   "Carrier_22_First_Duplicate_Carrier_Position" AT %QD1468 : DWord;
   "Carrier_22_Second_Duplicate_Carrier_Position" AT %QD1472 : DWord;
   "Carrier_22_CommandWord" AT %QW1476 : Word;
   "Carrier_22_Heartbeat" AT %Q1476.0 : Bool;
   "Carrier_22_Drive_Forward_Command" AT %Q1476.1 : Bool;
   "Carrier_22_Fault_Reset" AT %Q1476.2 : Bool;
   "Carrier_22_At_Command_Position" AT %Q1476.3 : Bool;
   "Carrier_22_Duplicate_Carrier_Fault" AT %Q1476.4 : Bool;
   "Carrier_22_Motion_On_Fault" AT %Q1476.5 : Bool;
   "Carrier_22_Motion_Off_Fault" AT %Q1476.6 : Bool;
   "Carrier_22_Carrier_Spacing_Fault" AT %Q1476.7 : Bool;
   "Carrier_23_Carrier_In_Zone" AT %QW1500 : Word;
   "Carrier_23_Carrier_Number_Echo" AT %QW1502 : Word;
   "Carrier_23_Carrier_Position_Echo" AT %QD1504 : DWord;
   "Carrier_23_Next_Carrier_Number" AT %QW1508 : Word;
   "Carrier_23_Next_Stop_Position" AT %QD1510 : DWord;
   "Carrier_23_Drive_Command_Speed" AT %QW1514 : Word;
   "Carrier_23_Duplicate_Carrier_Number" AT %QW1516 : Word;
   "Carrier_23_First_Duplicate_Carrier_Position" AT %QD1518 : DWord;
   "Carrier_23_Second_Duplicate_Carrier_Position" AT %QD1522 : DWord;
   "Carrier_23_CommandWord" AT %QW1526 : Word;
   "Carrier_23_Heartbeat" AT %Q1526.0 : Bool;
   "Carrier_23_Drive_Forward_Command" AT %Q1526.1 : Bool;
   "Carrier_23_Fault_Reset" AT %Q1526.2 : Bool;
   "Carrier_23_At_Command_Position" AT %Q1526.3 : Bool;
   "Carrier_23_Duplicate_Carrier_Fault" AT %Q1526.4 : Bool;
   "Carrier_23_Motion_On_Fault" AT %Q1526.5 : Bool;
   "Carrier_23_Motion_Off_Fault" AT %Q1526.6 : Bool;
   "Carrier_23_Carrier_Spacing_Fault" AT %Q1526.7 : Bool;
   "Carrier_24_Carrier_In_Zone" AT %QW1550 : Word;
   "Carrier_24_Carrier_Number_Echo" AT %QW1552 : Word;
   "Carrier_24_Carrier_Position_Echo" AT %QD1554 : DWord;
   "Carrier_24_Next_Carrier_Number" AT %QW1558 : Word;
   "Carrier_24_Next_Stop_Position" AT %QD1560 : DWord;
   "Carrier_24_Drive_Command_Speed" AT %QW1564 : Word;
   "Carrier_24_Duplicate_Carrier_Number" AT %QW1566 : Word;
   "Carrier_24_First_Duplicate_Carrier_Position" AT %QD1568 : DWord;
   "Carrier_24_Second_Duplicate_Carrier_Position" AT %QD1572 : DWord;
   "Carrier_24_CommandWord" AT %QW1576 : Word;
   "Carrier_24_Heartbeat" AT %Q1576.0 : Bool;
   "Carrier_24_Drive_Forward_Command" AT %Q1576.1 : Bool;
   "Carrier_24_Fault_Reset" AT %Q1576.2 : Bool;
   "Carrier_24_At_Command_Position" AT %Q1576.3 : Bool;
   "Carrier_24_Duplicate_Carrier_Fault" AT %Q1576.4 : Bool;
   "Carrier_24_Motion_On_Fault" AT %Q1576.5 : Bool;
   "Carrier_24_Motion_Off_Fault" AT %Q1576.6 : Bool;
   "Carrier_24_Carrier_Spacing_Fault" AT %Q1576.7 : Bool;
   "Carrier_25_Carrier_In_Zone" AT %QW1600 : Word;
   "Carrier_25_Carrier_Number_Echo" AT %QW1602 : Word;
   "Carrier_25_Carrier_Position_Echo" AT %QD1604 : DWord;
   "Carrier_25_Next_Carrier_Number" AT %QW1608 : Word;
   "Carrier_25_Next_Stop_Position" AT %QD1610 : DWord;
   "Carrier_25_Drive_Command_Speed" AT %QW1614 : Word;
   "Carrier_25_Duplicate_Carrier_Number" AT %QW1616 : Word;
   "Carrier_25_First_Duplicate_Carrier_Position" AT %QD1618 : DWord;
   "Carrier_25_Second_Duplicate_Carrier_Position" AT %QD1622 : DWord;
   "Carrier_25_CommandWord" AT %QW1626 : Word;
   "Carrier_25_Heartbeat" AT %Q1626.0 : Bool;
   "Carrier_25_Drive_Forward_Command" AT %Q1626.1 : Bool;
   "Carrier_25_Fault_Reset" AT %Q1626.2 : Bool;
   "Carrier_25_At_Command_Position" AT %Q1626.3 : Bool;
   "Carrier_25_Duplicate_Carrier_Fault" AT %Q1626.4 : Bool;
   "Carrier_25_Motion_On_Fault" AT %Q1626.5 : Bool;
   "Carrier_25_Motion_Off_Fault" AT %Q1626.6 : Bool;
   "Carrier_25_Carrier_Spacing_Fault" AT %Q1626.7 : Bool;
   "Carrier_26_Carrier_In_Zone" AT %QW1650 : Word;
   "Carrier_26_Carrier_Number_Echo" AT %QW1652 : Word;
   "Carrier_26_Carrier_Position_Echo" AT %QD1654 : DWord;
   "Carrier_26_Next_Carrier_Number" AT %QW1658 : Word;
   "Carrier_26_Next_Stop_Position" AT %QD1660 : DWord;
   "Carrier_26_Drive_Command_Speed" AT %QW1664 : Word;
   "Carrier_26_Duplicate_Carrier_Number" AT %QW1666 : Word;
   "Carrier_26_First_Duplicate_Carrier_Position" AT %QD1668 : DWord;
   "Carrier_26_Second_Duplicate_Carrier_Position" AT %QD1672 : DWord;
   "Carrier_26_CommandWord" AT %QW1676 : Word;
   "Carrier_26_Heartbeat" AT %Q1676.0 : Bool;
   "Carrier_26_Drive_Forward_Command" AT %Q1676.1 : Bool;
   "Carrier_26_Fault_Reset" AT %Q1676.2 : Bool;
   "Carrier_26_At_Command_Position" AT %Q1676.3 : Bool;
   "Carrier_26_Duplicate_Carrier_Fault" AT %Q1676.4 : Bool;
   "Carrier_26_Motion_On_Fault" AT %Q1676.5 : Bool;
   "Carrier_26_Motion_Off_Fault" AT %Q1676.6 : Bool;
   "Carrier_26_Carrier_Spacing_Fault" AT %Q1676.7 : Bool;
   "Carrier_27_Carrier_In_Zone" AT %QW1700 : Word;
   "Carrier_27_Carrier_Number_Echo" AT %QW1702 : Word;
   "Carrier_27_Carrier_Position_Echo" AT %QD1704 : DWord;
   "Carrier_27_Next_Carrier_Number" AT %QW1708 : Word;
   "Carrier_27_Next_Stop_Position" AT %QD1710 : DWord;
   "Carrier_27_Drive_Command_Speed" AT %QW1714 : Word;
   "Carrier_27_Duplicate_Carrier_Number" AT %QW1716 : Word;
   "Carrier_27_First_Duplicate_Carrier_Position" AT %QD1718 : DWord;
   "Carrier_27_Second_Duplicate_Carrier_Position" AT %QD1722 : DWord;
   "Carrier_27_CommandWord" AT %QW1726 : Word;
   "Carrier_27_Heartbeat" AT %Q1726.0 : Bool;
   "Carrier_27_Drive_Forward_Command" AT %Q1726.1 : Bool;
   "Carrier_27_Fault_Reset" AT %Q1726.2 : Bool;
   "Carrier_27_At_Command_Position" AT %Q1726.3 : Bool;
   "Carrier_27_Duplicate_Carrier_Fault" AT %Q1726.4 : Bool;
   "Carrier_27_Motion_On_Fault" AT %Q1726.5 : Bool;
   "Carrier_27_Motion_Off_Fault" AT %Q1726.6 : Bool;
   "Carrier_27_Carrier_Spacing_Fault" AT %Q1726.7 : Bool;
   "Carrier_28_Carrier_In_Zone" AT %QW1750 : Word;
   "Carrier_28_Carrier_Number_Echo" AT %QW1752 : Word;
   "Carrier_28_Carrier_Position_Echo" AT %QD1754 : DWord;
   "Carrier_28_Next_Carrier_Number" AT %QW1758 : Word;
   "Carrier_28_Next_Stop_Position" AT %QD1760 : DWord;
   "Carrier_28_Drive_Command_Speed" AT %QW1764 : Word;
   "Carrier_28_Duplicate_Carrier_Number" AT %QW1766 : Word;
   "Carrier_28_First_Duplicate_Carrier_Position" AT %QD1768 : DWord;
   "Carrier_28_Second_Duplicate_Carrier_Position" AT %QD1772 : DWord;
   "Carrier_28_CommandWord" AT %QW1776 : Word;
   "Carrier_28_Heartbeat" AT %Q1776.0 : Bool;
   "Carrier_28_Drive_Forward_Command" AT %Q1776.1 : Bool;
   "Carrier_28_Fault_Reset" AT %Q1776.2 : Bool;
   "Carrier_28_At_Command_Position" AT %Q1776.3 : Bool;
   "Carrier_28_Duplicate_Carrier_Fault" AT %Q1776.4 : Bool;
   "Carrier_28_Motion_On_Fault" AT %Q1776.5 : Bool;
   "Carrier_28_Motion_Off_Fault" AT %Q1776.6 : Bool;
   "Carrier_28_Carrier_Spacing_Fault" AT %Q1776.7 : Bool;
   "Carrier_29_Carrier_In_Zone" AT %QW1800 : Word;
   "Carrier_29_Carrier_Number_Echo" AT %QW1802 : Word;
   "Carrier_29_Carrier_Position_Echo" AT %QD1804 : DWord;
   "Carrier_29_Next_Carrier_Number" AT %QW1808 : Word;
   "Carrier_29_Next_Stop_Position" AT %QD1810 : DWord;
   "Carrier_29_Drive_Command_Speed" AT %QW1814 : Word;
   "Carrier_29_Duplicate_Carrier_Number" AT %QW1816 : Word;
   "Carrier_29_First_Duplicate_Carrier_Position" AT %QD1818 : DWord;
   "Carrier_29_Second_Duplicate_Carrier_Position" AT %QD1822 : DWord;
   "Carrier_29_CommandWord" AT %QW1826 : Word;
   "Carrier_29_Heartbeat" AT %Q1826.0 : Bool;
   "Carrier_29_Drive_Forward_Command" AT %Q1826.1 : Bool;
   "Carrier_29_Fault_Reset" AT %Q1826.2 : Bool;
   "Carrier_29_At_Command_Position" AT %Q1826.3 : Bool;
   "Carrier_29_Duplicate_Carrier_Fault" AT %Q1826.4 : Bool;
   "Carrier_29_Motion_On_Fault" AT %Q1826.5 : Bool;
   "Carrier_29_Motion_Off_Fault" AT %Q1826.6 : Bool;
   "Carrier_29_Carrier_Spacing_Fault" AT %Q1826.7 : Bool;
   "Carrier_30_Carrier_In_Zone" AT %QW1850 : Word;
   "Carrier_30_Carrier_Number_Echo" AT %QW1852 : Word;
   "Carrier_30_Carrier_Position_Echo" AT %QD1854 : DWord;
   "Carrier_30_Next_Carrier_Number" AT %QW1858 : Word;
   "Carrier_30_Next_Stop_Position" AT %QD1860 : DWord;
   "Carrier_30_Drive_Command_Speed" AT %QW1864 : Word;
   "Carrier_30_Duplicate_Carrier_Number" AT %QW1866 : Word;
   "Carrier_30_First_Duplicate_Carrier_Position" AT %QD1868 : DWord;
   "Carrier_30_Second_Duplicate_Carrier_Position" AT %QD1872 : DWord;
   "Carrier_30_CommandWord" AT %QW1876 : Word;
   "Carrier_30_Heartbeat" AT %Q1876.0 : Bool;
   "Carrier_30_Drive_Forward_Command" AT %Q1876.1 : Bool;
   "Carrier_30_Fault_Reset" AT %Q1876.2 : Bool;
   "Carrier_30_At_Command_Position" AT %Q1876.3 : Bool;
   "Carrier_30_Duplicate_Carrier_Fault" AT %Q1876.4 : Bool;
   "Carrier_30_Motion_On_Fault" AT %Q1876.5 : Bool;
   "Carrier_30_Motion_Off_Fault" AT %Q1876.6 : Bool;
   "Carrier_30_Carrier_Spacing_Fault" AT %Q1876.7 : Bool;
   "Carrier_31_Carrier_In_Zone" AT %QW1900 : Word;
   "Carrier_31_Carrier_Number_Echo" AT %QW1902 : Word;
   "Carrier_31_Carrier_Position_Echo" AT %QD1904 : DWord;
   "Carrier_31_Next_Carrier_Number" AT %QW1908 : Word;
   "Carrier_31_Next_Stop_Position" AT %QD1910 : DWord;
   "Carrier_31_Drive_Command_Speed" AT %QW1914 : Word;
   "Carrier_31_Duplicate_Carrier_Number" AT %QW1916 : Word;
   "Carrier_31_First_Duplicate_Carrier_Position" AT %QD1918 : DWord;
   "Carrier_31_Second_Duplicate_Carrier_Position" AT %QD1922 : DWord;
   "Carrier_31_CommandWord" AT %QW1926 : Word;
   "Carrier_31_Heartbeat" AT %Q1926.0 : Bool;
   "Carrier_31_Drive_Forward_Command" AT %Q1926.1 : Bool;
   "Carrier_31_Fault_Reset" AT %Q1926.2 : Bool;
   "Carrier_31_At_Command_Position" AT %Q1926.3 : Bool;
   "Carrier_31_Duplicate_Carrier_Fault" AT %Q1926.4 : Bool;
   "Carrier_31_Motion_On_Fault" AT %Q1926.5 : Bool;
   "Carrier_31_Motion_Off_Fault" AT %Q1926.6 : Bool;
   "Carrier_31_Carrier_Spacing_Fault" AT %Q1926.7 : Bool;
   "Carrier_32_Carrier_In_Zone" AT %QW1950 : Word;
   "Carrier_32_Carrier_Number_Echo" AT %QW1952 : Word;
   "Carrier_32_Carrier_Position_Echo" AT %QD1954 : DWord;
   "Carrier_32_Next_Carrier_Number" AT %QW1958 : Word;
   "Carrier_32_Next_Stop_Position" AT %QD1960 : DWord;
   "Carrier_32_Drive_Command_Speed" AT %QW1964 : Word;
   "Carrier_32_Duplicate_Carrier_Number" AT %QW1966 : Word;
   "Carrier_32_First_Duplicate_Carrier_Position" AT %QD1968 : DWord;
   "Carrier_32_Second_Duplicate_Carrier_Position" AT %QD1972 : DWord;
   "Carrier_32_CommandWord" AT %QW1976 : Word;
   "Carrier_32_Heartbeat" AT %Q1976.0 : Bool;
   "Carrier_32_Drive_Forward_Command" AT %Q1976.1 : Bool;
   "Carrier_32_Fault_Reset" AT %Q1976.2 : Bool;
   "Carrier_32_At_Command_Position" AT %Q1976.3 : Bool;
   "Carrier_32_Duplicate_Carrier_Fault" AT %Q1976.4 : Bool;
   "Carrier_32_Motion_On_Fault" AT %Q1976.5 : Bool;
   "Carrier_32_Motion_Off_Fault" AT %Q1976.6 : Bool;
   "Carrier_32_Carrier_Spacing_Fault" AT %Q1976.7 : Bool;
   "Carrier_33_Carrier_In_Zone" AT %QW2000 : Word;
   "Carrier_33_Carrier_Number_Echo" AT %QW2002 : Word;
   "Carrier_33_Carrier_Position_Echo" AT %QD2004 : DWord;
   "Carrier_33_Next_Carrier_Number" AT %QW2008 : Word;
   "Carrier_33_Next_Stop_Position" AT %QD2010 : DWord;
   "Carrier_33_Drive_Command_Speed" AT %QW2014 : Word;
   "Carrier_33_Duplicate_Carrier_Number" AT %QW2016 : Word;
   "Carrier_33_First_Duplicate_Carrier_Position" AT %QD2018 : DWord;
   "Carrier_33_Second_Duplicate_Carrier_Position" AT %QD2022 : DWord;
   "Carrier_33_CommandWord" AT %QW2026 : Word;
   "Carrier_33_Heartbeat" AT %Q2026.0 : Bool;
   "Carrier_33_Drive_Forward_Command" AT %Q2026.1 : Bool;
   "Carrier_33_Fault_Reset" AT %Q2026.2 : Bool;
   "Carrier_33_At_Command_Position" AT %Q2026.3 : Bool;
   "Carrier_33_Duplicate_Carrier_Fault" AT %Q2026.4 : Bool;
   "Carrier_33_Motion_On_Fault" AT %Q2026.5 : Bool;
   "Carrier_33_Motion_Off_Fault" AT %Q2026.6 : Bool;
   "Carrier_33_Carrier_Spacing_Fault" AT %Q2026.7 : Bool;
   "Carrier_34_Carrier_In_Zone" AT %QW2050 : Word;
   "Carrier_34_Carrier_Number_Echo" AT %QW2052 : Word;
   "Carrier_34_Carrier_Position_Echo" AT %QD2054 : DWord;
   "Carrier_34_Next_Carrier_Number" AT %QW2058 : Word;
   "Carrier_34_Next_Stop_Position" AT %QD2060 : DWord;
   "Carrier_34_Drive_Command_Speed" AT %QW2064 : Word;
   "Carrier_34_Duplicate_Carrier_Number" AT %QW2066 : Word;
   "Carrier_34_First_Duplicate_Carrier_Position" AT %QD2068 : DWord;
   "Carrier_34_Second_Duplicate_Carrier_Position" AT %QD2072 : DWord;
   "Carrier_34_CommandWord" AT %QW2076 : Word;
   "Carrier_34_Heartbeat" AT %Q2076.0 : Bool;
   "Carrier_34_Drive_Forward_Command" AT %Q2076.1 : Bool;
   "Carrier_34_Fault_Reset" AT %Q2076.2 : Bool;
   "Carrier_34_At_Command_Position" AT %Q2076.3 : Bool;
   "Carrier_34_Duplicate_Carrier_Fault" AT %Q2076.4 : Bool;
   "Carrier_34_Motion_On_Fault" AT %Q2076.5 : Bool;
   "Carrier_34_Motion_Off_Fault" AT %Q2076.6 : Bool;
   "Carrier_34_Carrier_Spacing_Fault" AT %Q2076.7 : Bool;
   "Carrier_35_Carrier_In_Zone" AT %QW2100 : Word;
   "Carrier_35_Carrier_Number_Echo" AT %QW2102 : Word;
   "Carrier_35_Carrier_Position_Echo" AT %QD2104 : DWord;
   "Carrier_35_Next_Carrier_Number" AT %QW2108 : Word;
   "Carrier_35_Next_Stop_Position" AT %QD2110 : DWord;
   "Carrier_35_Drive_Command_Speed" AT %QW2114 : Word;
   "Carrier_35_Duplicate_Carrier_Number" AT %QW2116 : Word;
   "Carrier_35_First_Duplicate_Carrier_Position" AT %QD2118 : DWord;
   "Carrier_35_Second_Duplicate_Carrier_Position" AT %QD2122 : DWord;
   "Carrier_35_CommandWord" AT %QW2126 : Word;
   "Carrier_35_Heartbeat" AT %Q2126.0 : Bool;
   "Carrier_35_Drive_Forward_Command" AT %Q2126.1 : Bool;
   "Carrier_35_Fault_Reset" AT %Q2126.2 : Bool;
   "Carrier_35_At_Command_Position" AT %Q2126.3 : Bool;
   "Carrier_35_Duplicate_Carrier_Fault" AT %Q2126.4 : Bool;
   "Carrier_35_Motion_On_Fault" AT %Q2126.5 : Bool;
   "Carrier_35_Motion_Off_Fault" AT %Q2126.6 : Bool;
   "Carrier_35_Carrier_Spacing_Fault" AT %Q2126.7 : Bool;
   "Carrier_36_Carrier_In_Zone" AT %QW2150 : Word;
   "Carrier_36_Carrier_Number_Echo" AT %QW2152 : Word;
   "Carrier_36_Carrier_Position_Echo" AT %QD2154 : DWord;
   "Carrier_36_Next_Carrier_Number" AT %QW2158 : Word;
   "Carrier_36_Next_Stop_Position" AT %QD2160 : DWord;
   "Carrier_36_Drive_Command_Speed" AT %QW2164 : Word;
   "Carrier_36_Duplicate_Carrier_Number" AT %QW2166 : Word;
   "Carrier_36_First_Duplicate_Carrier_Position" AT %QD2168 : DWord;
   "Carrier_36_Second_Duplicate_Carrier_Position" AT %QD2172 : DWord;
   "Carrier_36_CommandWord" AT %QW2176 : Word;
   "Carrier_36_Heartbeat" AT %Q2176.0 : Bool;
   "Carrier_36_Drive_Forward_Command" AT %Q2176.1 : Bool;
   "Carrier_36_Fault_Reset" AT %Q2176.2 : Bool;
   "Carrier_36_At_Command_Position" AT %Q2176.3 : Bool;
   "Carrier_36_Duplicate_Carrier_Fault" AT %Q2176.4 : Bool;
   "Carrier_36_Motion_On_Fault" AT %Q2176.5 : Bool;
   "Carrier_36_Motion_Off_Fault" AT %Q2176.6 : Bool;
   "Carrier_36_Carrier_Spacing_Fault" AT %Q2176.7 : Bool;
   "Carrier_37_Carrier_In_Zone" AT %QW2200 : Word;
   "Carrier_37_Carrier_Number_Echo" AT %QW2202 : Word;
   "Carrier_37_Carrier_Position_Echo" AT %QD2204 : DWord;
   "Carrier_37_Next_Carrier_Number" AT %QW2208 : Word;
   "Carrier_37_Next_Stop_Position" AT %QD2210 : DWord;
   "Carrier_37_Drive_Command_Speed" AT %QW2214 : Word;
   "Carrier_37_Duplicate_Carrier_Number" AT %QW2216 : Word;
   "Carrier_37_First_Duplicate_Carrier_Position" AT %QD2218 : DWord;
   "Carrier_37_Second_Duplicate_Carrier_Position" AT %QD2222 : DWord;
   "Carrier_37_CommandWord" AT %QW2226 : Word;
   "Carrier_37_Heartbeat" AT %Q2226.0 : Bool;
   "Carrier_37_Drive_Forward_Command" AT %Q2226.1 : Bool;
   "Carrier_37_Fault_Reset" AT %Q2226.2 : Bool;
   "Carrier_37_At_Command_Position" AT %Q2226.3 : Bool;
   "Carrier_37_Duplicate_Carrier_Fault" AT %Q2226.4 : Bool;
   "Carrier_37_Motion_On_Fault" AT %Q2226.5 : Bool;
   "Carrier_37_Motion_Off_Fault" AT %Q2226.6 : Bool;
   "Carrier_37_Carrier_Spacing_Fault" AT %Q2226.7 : Bool;
   "Carrier_38_Carrier_In_Zone" AT %QW2250 : Word;
   "Carrier_38_Carrier_Number_Echo" AT %QW2252 : Word;
   "Carrier_38_Carrier_Position_Echo" AT %QD2254 : DWord;
   "Carrier_38_Next_Carrier_Number" AT %QW2258 : Word;
   "Carrier_38_Next_Stop_Position" AT %QD2260 : DWord;
   "Carrier_38_Drive_Command_Speed" AT %QW2264 : Word;
   "Carrier_38_Duplicate_Carrier_Number" AT %QW2266 : Word;
   "Carrier_38_First_Duplicate_Carrier_Position" AT %QD2268 : DWord;
   "Carrier_38_Second_Duplicate_Carrier_Position" AT %QD2272 : DWord;
   "Carrier_38_CommandWord" AT %QW2276 : Word;
   "Carrier_38_Heartbeat" AT %Q2276.0 : Bool;
   "Carrier_38_Drive_Forward_Command" AT %Q2276.1 : Bool;
   "Carrier_38_Fault_Reset" AT %Q2276.2 : Bool;
   "Carrier_38_At_Command_Position" AT %Q2276.3 : Bool;
   "Carrier_38_Duplicate_Carrier_Fault" AT %Q2276.4 : Bool;
   "Carrier_38_Motion_On_Fault" AT %Q2276.5 : Bool;
   "Carrier_38_Motion_Off_Fault" AT %Q2276.6 : Bool;
   "Carrier_38_Carrier_Spacing_Fault" AT %Q2276.7 : Bool;
   "Carrier_39_Carrier_In_Zone" AT %QW2300 : Word;
   "Carrier_39_Carrier_Number_Echo" AT %QW2302 : Word;
   "Carrier_39_Carrier_Position_Echo" AT %QD2304 : DWord;
   "Carrier_39_Next_Carrier_Number" AT %QW2308 : Word;
   "Carrier_39_Next_Stop_Position" AT %QD2310 : DWord;
   "Carrier_39_Drive_Command_Speed" AT %QW2314 : Word;
   "Carrier_39_Duplicate_Carrier_Number" AT %QW2316 : Word;
   "Carrier_39_First_Duplicate_Carrier_Position" AT %QD2318 : DWord;
   "Carrier_39_Second_Duplicate_Carrier_Position" AT %QD2322 : DWord;
   "Carrier_39_CommandWord" AT %QW2326 : Word;
   "Carrier_39_Heartbeat" AT %Q2326.0 : Bool;
   "Carrier_39_Drive_Forward_Command" AT %Q2326.1 : Bool;
   "Carrier_39_Fault_Reset" AT %Q2326.2 : Bool;
   "Carrier_39_At_Command_Position" AT %Q2326.3 : Bool;
   "Carrier_39_Duplicate_Carrier_Fault" AT %Q2326.4 : Bool;
   "Carrier_39_Motion_On_Fault" AT %Q2326.5 : Bool;
   "Carrier_39_Motion_Off_Fault" AT %Q2326.6 : Bool;
   "Carrier_39_Carrier_Spacing_Fault" AT %Q2326.7 : Bool;
   "Carrier_40_Carrier_In_Zone" AT %QW2350 : Word;
   "Carrier_40_Carrier_Number_Echo" AT %QW2352 : Word;
   "Carrier_40_Carrier_Position_Echo" AT %QD2354 : DWord;
   "Carrier_40_Next_Carrier_Number" AT %QW2358 : Word;
   "Carrier_40_Next_Stop_Position" AT %QD2360 : DWord;
   "Carrier_40_Drive_Command_Speed" AT %QW2364 : Word;
   "Carrier_40_Duplicate_Carrier_Number" AT %QW2366 : Word;
   "Carrier_40_First_Duplicate_Carrier_Position" AT %QD2368 : DWord;
   "Carrier_40_Second_Duplicate_Carrier_Position" AT %QD2372 : DWord;
   "Carrier_40_CommandWord" AT %QW2376 : Word;
   "Carrier_40_Heartbeat" AT %Q2376.0 : Bool;
   "Carrier_40_Drive_Forward_Command" AT %Q2376.1 : Bool;
   "Carrier_40_Fault_Reset" AT %Q2376.2 : Bool;
   "Carrier_40_At_Command_Position" AT %Q2376.3 : Bool;
   "Carrier_40_Duplicate_Carrier_Fault" AT %Q2376.4 : Bool;
   "Carrier_40_Motion_On_Fault" AT %Q2376.5 : Bool;
   "Carrier_40_Motion_Off_Fault" AT %Q2376.6 : Bool;
   "Carrier_40_Carrier_Spacing_Fault" AT %Q2376.7 : Bool;
   "Carrier_41_Carrier_In_Zone" AT %QW2400 : Word;
   "Carrier_41_Carrier_Number_Echo" AT %QW2402 : Word;
   "Carrier_41_Carrier_Position_Echo" AT %QD2404 : DWord;
   "Carrier_41_Next_Carrier_Number" AT %QW2408 : Word;
   "Carrier_41_Next_Stop_Position" AT %QD2410 : DWord;
   "Carrier_41_Drive_Command_Speed" AT %QW2414 : Word;
   "Carrier_41_Duplicate_Carrier_Number" AT %QW2416 : Word;
   "Carrier_41_First_Duplicate_Carrier_Position" AT %QD2418 : DWord;
   "Carrier_41_Second_Duplicate_Carrier_Position" AT %QD2422 : DWord;
   "Carrier_41_CommandWord" AT %QW2426 : Word;
   "Carrier_41_Heartbeat" AT %Q2426.0 : Bool;
   "Carrier_41_Drive_Forward_Command" AT %Q2426.1 : Bool;
   "Carrier_41_Fault_Reset" AT %Q2426.2 : Bool;
   "Carrier_41_At_Command_Position" AT %Q2426.3 : Bool;
   "Carrier_41_Duplicate_Carrier_Fault" AT %Q2426.4 : Bool;
   "Carrier_41_Motion_On_Fault" AT %Q2426.5 : Bool;
   "Carrier_41_Motion_Off_Fault" AT %Q2426.6 : Bool;
   "Carrier_41_Carrier_Spacing_Fault" AT %Q2426.7 : Bool;
   "Carrier_42_Carrier_In_Zone" AT %QW2450 : Word;
   "Carrier_42_Carrier_Number_Echo" AT %QW2452 : Word;
   "Carrier_42_Carrier_Position_Echo" AT %QD2454 : DWord;
   "Carrier_42_Next_Carrier_Number" AT %QW2458 : Word;
   "Carrier_42_Next_Stop_Position" AT %QD2460 : DWord;
   "Carrier_42_Drive_Command_Speed" AT %QW2464 : Word;
   "Carrier_42_Duplicate_Carrier_Number" AT %QW2466 : Word;
   "Carrier_42_First_Duplicate_Carrier_Position" AT %QD2468 : DWord;
   "Carrier_42_Second_Duplicate_Carrier_Position" AT %QD2472 : DWord;
   "Carrier_42_CommandWord" AT %QW2476 : Word;
   "Carrier_42_Heartbeat" AT %Q2476.0 : Bool;
   "Carrier_42_Drive_Forward_Command" AT %Q2476.1 : Bool;
   "Carrier_42_Fault_Reset" AT %Q2476.2 : Bool;
   "Carrier_42_At_Command_Position" AT %Q2476.3 : Bool;
   "Carrier_42_Duplicate_Carrier_Fault" AT %Q2476.4 : Bool;
   "Carrier_42_Motion_On_Fault" AT %Q2476.5 : Bool;
   "Carrier_42_Motion_Off_Fault" AT %Q2476.6 : Bool;
   "Carrier_42_Carrier_Spacing_Fault" AT %Q2476.7 : Bool;
   "Carrier_43_Carrier_In_Zone" AT %QW2500 : Word;
   "Carrier_43_Carrier_Number_Echo" AT %QW2502 : Word;
   "Carrier_43_Carrier_Position_Echo" AT %QD2504 : DWord;
   "Carrier_43_Next_Carrier_Number" AT %QW2508 : Word;
   "Carrier_43_Next_Stop_Position" AT %QD2510 : DWord;
   "Carrier_43_Drive_Command_Speed" AT %QW2514 : Word;
   "Carrier_43_Duplicate_Carrier_Number" AT %QW2516 : Word;
   "Carrier_43_First_Duplicate_Carrier_Position" AT %QD2518 : DWord;
   "Carrier_43_Second_Duplicate_Carrier_Position" AT %QD2522 : DWord;
   "Carrier_43_CommandWord" AT %QW2526 : Word;
   "Carrier_43_Heartbeat" AT %Q2526.0 : Bool;
   "Carrier_43_Drive_Forward_Command" AT %Q2526.1 : Bool;
   "Carrier_43_Fault_Reset" AT %Q2526.2 : Bool;
   "Carrier_43_At_Command_Position" AT %Q2526.3 : Bool;
   "Carrier_43_Duplicate_Carrier_Fault" AT %Q2526.4 : Bool;
   "Carrier_43_Motion_On_Fault" AT %Q2526.5 : Bool;
   "Carrier_43_Motion_Off_Fault" AT %Q2526.6 : Bool;
   "Carrier_43_Carrier_Spacing_Fault" AT %Q2526.7 : Bool;
   "Carrier_44_Carrier_In_Zone" AT %QW2550 : Word;
   "Carrier_44_Carrier_Number_Echo" AT %QW2552 : Word;
   "Carrier_44_Carrier_Position_Echo" AT %QD2554 : DWord;
   "Carrier_44_Next_Carrier_Number" AT %QW2558 : Word;
   "Carrier_44_Next_Stop_Position" AT %QD2560 : DWord;
   "Carrier_44_Drive_Command_Speed" AT %QW2564 : Word;
   "Carrier_44_Duplicate_Carrier_Number" AT %QW2566 : Word;
   "Carrier_44_First_Duplicate_Carrier_Position" AT %QD2568 : DWord;
   "Carrier_44_Second_Duplicate_Carrier_Position" AT %QD2572 : DWord;
   "Carrier_44_CommandWord" AT %QW2576 : Word;
   "Carrier_44_Heartbeat" AT %Q2576.0 : Bool;
   "Carrier_44_Drive_Forward_Command" AT %Q2576.1 : Bool;
   "Carrier_44_Fault_Reset" AT %Q2576.2 : Bool;
   "Carrier_44_At_Command_Position" AT %Q2576.3 : Bool;
   "Carrier_44_Duplicate_Carrier_Fault" AT %Q2576.4 : Bool;
   "Carrier_44_Motion_On_Fault" AT %Q2576.5 : Bool;
   "Carrier_44_Motion_Off_Fault" AT %Q2576.6 : Bool;
   "Carrier_44_Carrier_Spacing_Fault" AT %Q2576.7 : Bool;
   "Carrier_45_Carrier_In_Zone" AT %QW2600 : Word;
   "Carrier_45_Carrier_Number_Echo" AT %QW2602 : Word;
   "Carrier_45_Carrier_Position_Echo" AT %QD2604 : DWord;
   "Carrier_45_Next_Carrier_Number" AT %QW2608 : Word;
   "Carrier_45_Next_Stop_Position" AT %QD2610 : DWord;
   "Carrier_45_Drive_Command_Speed" AT %QW2614 : Word;
   "Carrier_45_Duplicate_Carrier_Number" AT %QW2616 : Word;
   "Carrier_45_First_Duplicate_Carrier_Position" AT %QD2618 : DWord;
   "Carrier_45_Second_Duplicate_Carrier_Position" AT %QD2622 : DWord;
   "Carrier_45_CommandWord" AT %QW2626 : Word;
   "Carrier_45_Heartbeat" AT %Q2626.0 : Bool;
   "Carrier_45_Drive_Forward_Command" AT %Q2626.1 : Bool;
   "Carrier_45_Fault_Reset" AT %Q2626.2 : Bool;
   "Carrier_45_At_Command_Position" AT %Q2626.3 : Bool;
   "Carrier_45_Duplicate_Carrier_Fault" AT %Q2626.4 : Bool;
   "Carrier_45_Motion_On_Fault" AT %Q2626.5 : Bool;
   "Carrier_45_Motion_Off_Fault" AT %Q2626.6 : Bool;
   "Carrier_45_Carrier_Spacing_Fault" AT %Q2626.7 : Bool;
   "Carrier_46_Carrier_In_Zone" AT %QW2650 : Word;
   "Carrier_46_Carrier_Number_Echo" AT %QW2652 : Word;
   "Carrier_46_Carrier_Position_Echo" AT %QD2654 : DWord;
   "Carrier_46_Next_Carrier_Number" AT %QW2658 : Word;
   "Carrier_46_Next_Stop_Position" AT %QD2660 : DWord;
   "Carrier_46_Drive_Command_Speed" AT %QW2664 : Word;
   "Carrier_46_Duplicate_Carrier_Number" AT %QW2666 : Word;
   "Carrier_46_First_Duplicate_Carrier_Position" AT %QD2668 : DWord;
   "Carrier_46_Second_Duplicate_Carrier_Position" AT %QD2672 : DWord;
   "Carrier_46_CommandWord" AT %QW2676 : Word;
   "Carrier_46_Heartbeat" AT %Q2676.0 : Bool;
   "Carrier_46_Drive_Forward_Command" AT %Q2676.1 : Bool;
   "Carrier_46_Fault_Reset" AT %Q2676.2 : Bool;
   "Carrier_46_At_Command_Position" AT %Q2676.3 : Bool;
   "Carrier_46_Duplicate_Carrier_Fault" AT %Q2676.4 : Bool;
   "Carrier_46_Motion_On_Fault" AT %Q2676.5 : Bool;
   "Carrier_46_Motion_Off_Fault" AT %Q2676.6 : Bool;
   "Carrier_46_Carrier_Spacing_Fault" AT %Q2676.7 : Bool;
   "Carrier_47_Carrier_In_Zone" AT %QW2700 : Word;
   "Carrier_47_Carrier_Number_Echo" AT %QW2702 : Word;
   "Carrier_47_Carrier_Position_Echo" AT %QD2704 : DWord;
   "Carrier_47_Next_Carrier_Number" AT %QW2708 : Word;
   "Carrier_47_Next_Stop_Position" AT %QD2710 : DWord;
   "Carrier_47_Drive_Command_Speed" AT %QW2714 : Word;
   "Carrier_47_Duplicate_Carrier_Number" AT %QW2716 : Word;
   "Carrier_47_First_Duplicate_Carrier_Position" AT %QD2718 : DWord;
   "Carrier_47_Second_Duplicate_Carrier_Position" AT %QD2722 : DWord;
   "Carrier_47_CommandWord" AT %QW2726 : Word;
   "Carrier_47_Heartbeat" AT %Q2726.0 : Bool;
   "Carrier_47_Drive_Forward_Command" AT %Q2726.1 : Bool;
   "Carrier_47_Fault_Reset" AT %Q2726.2 : Bool;
   "Carrier_47_At_Command_Position" AT %Q2726.3 : Bool;
   "Carrier_47_Duplicate_Carrier_Fault" AT %Q2726.4 : Bool;
   "Carrier_47_Motion_On_Fault" AT %Q2726.5 : Bool;
   "Carrier_47_Motion_Off_Fault" AT %Q2726.6 : Bool;
   "Carrier_47_Carrier_Spacing_Fault" AT %Q2726.7 : Bool;
   "Carrier_48_Carrier_In_Zone" AT %QW2750 : Word;
   "Carrier_48_Carrier_Number_Echo" AT %QW2752 : Word;
   "Carrier_48_Carrier_Position_Echo" AT %QD2754 : DWord;
   "Carrier_48_Next_Carrier_Number" AT %QW2758 : Word;
   "Carrier_48_Next_Stop_Position" AT %QD2760 : DWord;
   "Carrier_48_Drive_Command_Speed" AT %QW2764 : Word;
   "Carrier_48_Duplicate_Carrier_Number" AT %QW2766 : Word;
   "Carrier_48_First_Duplicate_Carrier_Position" AT %QD2768 : DWord;
   "Carrier_48_Second_Duplicate_Carrier_Position" AT %QD2772 : DWord;
   "Carrier_48_CommandWord" AT %QW2776 : Word;
   "Carrier_48_Heartbeat" AT %Q2776.0 : Bool;
   "Carrier_48_Drive_Forward_Command" AT %Q2776.1 : Bool;
   "Carrier_48_Fault_Reset" AT %Q2776.2 : Bool;
   "Carrier_48_At_Command_Position" AT %Q2776.3 : Bool;
   "Carrier_48_Duplicate_Carrier_Fault" AT %Q2776.4 : Bool;
   "Carrier_48_Motion_On_Fault" AT %Q2776.5 : Bool;
   "Carrier_48_Motion_Off_Fault" AT %Q2776.6 : Bool;
   "Carrier_48_Carrier_Spacing_Fault" AT %Q2776.7 : Bool;
   "Carrier_49_Carrier_In_Zone" AT %QW2800 : Word;
   "Carrier_49_Carrier_Number_Echo" AT %QW2802 : Word;
   "Carrier_49_Carrier_Position_Echo" AT %QD2804 : DWord;
   "Carrier_49_Next_Carrier_Number" AT %QW2808 : Word;
   "Carrier_49_Next_Stop_Position" AT %QD2810 : DWord;
   "Carrier_49_Drive_Command_Speed" AT %QW2814 : Word;
   "Carrier_49_Duplicate_Carrier_Number" AT %QW2816 : Word;
   "Carrier_49_First_Duplicate_Carrier_Position" AT %QD2818 : DWord;
   "Carrier_49_Second_Duplicate_Carrier_Position" AT %QD2822 : DWord;
   "Carrier_49_CommandWord" AT %QW2826 : Word;
   "Carrier_49_Heartbeat" AT %Q2826.0 : Bool;
   "Carrier_49_Drive_Forward_Command" AT %Q2826.1 : Bool;
   "Carrier_49_Fault_Reset" AT %Q2826.2 : Bool;
   "Carrier_49_At_Command_Position" AT %Q2826.3 : Bool;
   "Carrier_49_Duplicate_Carrier_Fault" AT %Q2826.4 : Bool;
   "Carrier_49_Motion_On_Fault" AT %Q2826.5 : Bool;
   "Carrier_49_Motion_Off_Fault" AT %Q2826.6 : Bool;
   "Carrier_49_Carrier_Spacing_Fault" AT %Q2826.7 : Bool;
   "Carrier_50_Carrier_In_Zone" AT %QW2850 : Word;
   "Carrier_50_Carrier_Number_Echo" AT %QW2852 : Word;
   "Carrier_50_Carrier_Position_Echo" AT %QD2854 : DWord;
   "Carrier_50_Next_Carrier_Number" AT %QW2858 : Word;
   "Carrier_50_Next_Stop_Position" AT %QD2860 : DWord;
   "Carrier_50_Drive_Command_Speed" AT %QW2864 : Word;
   "Carrier_50_Duplicate_Carrier_Number" AT %QW2866 : Word;
   "Carrier_50_First_Duplicate_Carrier_Position" AT %QD2868 : DWord;
   "Carrier_50_Second_Duplicate_Carrier_Position" AT %QD2872 : DWord;
   "Carrier_50_CommandWord" AT %QW2876 : Word;
   "Carrier_50_Heartbeat" AT %Q2876.0 : Bool;
   "Carrier_50_Drive_Forward_Command" AT %Q2876.1 : Bool;
   "Carrier_50_Fault_Reset" AT %Q2876.2 : Bool;
   "Carrier_50_At_Command_Position" AT %Q2876.3 : Bool;
   "Carrier_50_Duplicate_Carrier_Fault" AT %Q2876.4 : Bool;
   "Carrier_50_Motion_On_Fault" AT %Q2876.5 : Bool;
   "Carrier_50_Motion_Off_Fault" AT %Q2876.6 : Bool;
   "Carrier_50_Carrier_Spacing_Fault" AT %Q2876.7 : Bool;
   "Carrier_51_Carrier_In_Zone" AT %QW2900 : Word;
   "Carrier_51_Carrier_Number_Echo" AT %QW2902 : Word;
   "Carrier_51_Carrier_Position_Echo" AT %QD2904 : DWord;
   "Carrier_51_Next_Carrier_Number" AT %QW2908 : Word;
   "Carrier_51_Next_Stop_Position" AT %QD2910 : DWord;
   "Carrier_51_Drive_Command_Speed" AT %QW2914 : Word;
   "Carrier_51_Duplicate_Carrier_Number" AT %QW2916 : Word;
   "Carrier_51_First_Duplicate_Carrier_Position" AT %QD2918 : DWord;
   "Carrier_51_Second_Duplicate_Carrier_Position" AT %QD2922 : DWord;
   "Carrier_51_CommandWord" AT %QW2926 : Word;
   "Carrier_51_Heartbeat" AT %Q2926.0 : Bool;
   "Carrier_51_Drive_Forward_Command" AT %Q2926.1 : Bool;
   "Carrier_51_Fault_Reset" AT %Q2926.2 : Bool;
   "Carrier_51_At_Command_Position" AT %Q2926.3 : Bool;
   "Carrier_51_Duplicate_Carrier_Fault" AT %Q2926.4 : Bool;
   "Carrier_51_Motion_On_Fault" AT %Q2926.5 : Bool;
   "Carrier_51_Motion_Off_Fault" AT %Q2926.6 : Bool;
   "Carrier_51_Carrier_Spacing_Fault" AT %Q2926.7 : Bool;
   "Carrier_52_Carrier_In_Zone" AT %QW2950 : Word;
   "Carrier_52_Carrier_Number_Echo" AT %QW2952 : Word;
   "Carrier_52_Carrier_Position_Echo" AT %QD2954 : DWord;
   "Carrier_52_Next_Carrier_Number" AT %QW2958 : Word;
   "Carrier_52_Next_Stop_Position" AT %QD2960 : DWord;
   "Carrier_52_Drive_Command_Speed" AT %QW2964 : Word;
   "Carrier_52_Duplicate_Carrier_Number" AT %QW2966 : Word;
   "Carrier_52_First_Duplicate_Carrier_Position" AT %QD2968 : DWord;
   "Carrier_52_Second_Duplicate_Carrier_Position" AT %QD2972 : DWord;
   "Carrier_52_CommandWord" AT %QW2976 : Word;
   "Carrier_52_Heartbeat" AT %Q2976.0 : Bool;
   "Carrier_52_Drive_Forward_Command" AT %Q2976.1 : Bool;
   "Carrier_52_Fault_Reset" AT %Q2976.2 : Bool;
   "Carrier_52_At_Command_Position" AT %Q2976.3 : Bool;
   "Carrier_52_Duplicate_Carrier_Fault" AT %Q2976.4 : Bool;
   "Carrier_52_Motion_On_Fault" AT %Q2976.5 : Bool;
   "Carrier_52_Motion_Off_Fault" AT %Q2976.6 : Bool;
   "Carrier_52_Carrier_Spacing_Fault" AT %Q2976.7 : Bool;
   "Carrier_53_Carrier_In_Zone" AT %QW3000 : Word;
   "Carrier_53_Carrier_Number_Echo" AT %QW3002 : Word;
   "Carrier_53_Carrier_Position_Echo" AT %QD3004 : DWord;
   "Carrier_53_Next_Carrier_Number" AT %QW3008 : Word;
   "Carrier_53_Next_Stop_Position" AT %QD3010 : DWord;
   "Carrier_53_Drive_Command_Speed" AT %QW3014 : Word;
   "Carrier_53_Duplicate_Carrier_Number" AT %QW3016 : Word;
   "Carrier_53_First_Duplicate_Carrier_Position" AT %QD3018 : DWord;
   "Carrier_53_Second_Duplicate_Carrier_Position" AT %QD3022 : DWord;
   "Carrier_53_CommandWord" AT %QW3026 : Word;
   "Carrier_53_Heartbeat" AT %Q3026.0 : Bool;
   "Carrier_53_Drive_Forward_Command" AT %Q3026.1 : Bool;
   "Carrier_53_Fault_Reset" AT %Q3026.2 : Bool;
   "Carrier_53_At_Command_Position" AT %Q3026.3 : Bool;
   "Carrier_53_Duplicate_Carrier_Fault" AT %Q3026.4 : Bool;
   "Carrier_53_Motion_On_Fault" AT %Q3026.5 : Bool;
   "Carrier_53_Motion_Off_Fault" AT %Q3026.6 : Bool;
   "Carrier_53_Carrier_Spacing_Fault" AT %Q3026.7 : Bool;
   "Carrier_54_Carrier_In_Zone" AT %QW3050 : Word;
   "Carrier_54_Carrier_Number_Echo" AT %QW3052 : Word;
   "Carrier_54_Carrier_Position_Echo" AT %QD3054 : DWord;
   "Carrier_54_Next_Carrier_Number" AT %QW3058 : Word;
   "Carrier_54_Next_Stop_Position" AT %QD3060 : DWord;
   "Carrier_54_Drive_Command_Speed" AT %QW3064 : Word;
   "Carrier_54_Duplicate_Carrier_Number" AT %QW3066 : Word;
   "Carrier_54_First_Duplicate_Carrier_Position" AT %QD3068 : DWord;
   "Carrier_54_Second_Duplicate_Carrier_Position" AT %QD3072 : DWord;
   "Carrier_54_CommandWord" AT %QW3076 : Word;
   "Carrier_54_Heartbeat" AT %Q3076.0 : Bool;
   "Carrier_54_Drive_Forward_Command" AT %Q3076.1 : Bool;
   "Carrier_54_Fault_Reset" AT %Q3076.2 : Bool;
   "Carrier_54_At_Command_Position" AT %Q3076.3 : Bool;
   "Carrier_54_Duplicate_Carrier_Fault" AT %Q3076.4 : Bool;
   "Carrier_54_Motion_On_Fault" AT %Q3076.5 : Bool;
   "Carrier_54_Motion_Off_Fault" AT %Q3076.6 : Bool;
   "Carrier_54_Carrier_Spacing_Fault" AT %Q3076.7 : Bool;
   "Carrier_55_Carrier_In_Zone" AT %QW3100 : Word;